VERSION : 0.1
   VAR_INPUT
      digits : String;
   END_VAR
   VAR_TEMP
      _characters : Array[0..#CHAR_COUNT] of Char;
      _count : DInt;
      _i : Int;
      _length : Int;
      _character_count : Int;
      _return : DInt;
      _temp : Bool;
   END_VAR
   VAR CONSTANT
      ASCII_OFFSET : DInt := 16#30;
      BLANK : Time;
      CHAR_COUNT : Int := 9;
      MS_PER_SEC : DInt := 1_000;
   END_VAR
BEGIN
   REGION "EXIT ON NO INPUT"
       IF #digits = '' THEN
           #"Timer.Digits_as_String_to_Seconds" := #BLANK;
           RETURN;
       END_IF;
   END_REGION


   REGION "EXPLODE"
       Strg_TO_Chars(Strg := #digits,
                     pChars := 0,
                     Cnt => #_count,
                     Chars := #_characters);
       #_length := UDINT_TO_INT("Array.Any.Length"(#_characters)) - 1;
   END_REGION


   REGION "COUNT"
       #_character_count := "Array.Char.Search"(array := #_characters, search_term := ' ') - 1;
   END_REGION


   REGION "VALIDATE"
       FOR #_i := 0 TO #_character_count DO
           IF NOT "Char.Is_Numeric"(#_characters[#_i]) THEN
               #"Timer.Digits_as_String_to_Seconds" := #BLANK;
               RETURN;
           END_IF;
       END_FOR;
   END_REGION


   #"Timer.Digits_as_String_to_Seconds" := STRING_TO_DINT(#digits) * #MS_PER_SEC;
END_FUNCTION

FUNCTION "Timer.Digits_as_String_to_Minutes" : Time   // FC267, SCL
{ S7_Optimized_Access := 'TRUE' }
VERSION : 0.1
   VAR_INPUT
      digits : String;
   END_VAR
   VAR CONSTANT
      SECONDS_PER_MINUTE : Int := 60;
   END_VAR
BEGIN
   #"Timer.Digits_as_String_to_Minutes" := #SECONDS_PER_MINUTE * TIME_TO_DINT("Timer.Digits_as_String_to_Seconds"(#digits));
END_FUNCTION

FUNCTION "Timer.Digits_as_String_to_Hours" : Time   // FC269, SCL
{ S7_Optimized_Access := 'TRUE' }
VERSION : 0.1
   VAR_INPUT
      digits : String;
   END_VAR
   VAR CONSTANT
      SECONDS_PER_HOUR : Int := 3_600;
   END_VAR
BEGIN
   #"Timer.Digits_as_String_to_Hours" := #SECONDS_PER_HOUR * TIME_TO_DINT("Timer.Digits_as_String_to_Seconds"(#digits));
END_FUNCTION

// folder: Utilities/UInt

FUNCTION "UInt.Value_Change" : Bool   // FC183, SCL
{ S7_Optimized_Access := 'TRUE' }
VERSION : 0.1
   VAR_INPUT
      value : UInt;
      old_value : UInt;
   END_VAR
BEGIN
   #"UInt.Value_Change" := #value <> #old_value;
END_FUNCTION

// folder: Utilities/USInt

FUNCTION_BLOCK "USInt.State_change"   // FB58, SCL
{ S7_Optimized_Access := 'TRUE' }
VERSION : 0.1
   VAR_INPUT
      value : USInt;
   END_VAR
   VAR_IN_OUT
      get_usint : "State Changes: USInt";
   END_VAR
   VAR
      old_value : USInt;
   END_VAR
   VAR_TEMP
      _return : "State Changes: USInt";
   END_VAR
BEGIN
   REGION "BUFFER IN"
       #_return := #get_usint;
   END_REGION


   REGION "MAP"
       IF #value <> #old_value THEN
           #_return.actual := #value;
       END_IF;
       #_return.rising := "USInt.Rising_Edge"(value := #value,
                                              old_value := #old_value);
       #_return.falling := "USInt.Falling_Edge"(value := #value,
                                                old_value := #old_value);
   END_REGION


   REGION "SAVE OLD VALUE"
       #old_value := #_return.actual;
   END_REGION


   REGION "RETURN" 
       #get_usint := #_return;
   END_REGION
END_FUNCTION_BLOCK

FUNCTION "USInt.Value_Change" : Bool   // FC181, SCL
{ S7_Optimized_Access := 'TRUE' }
VERSION : 0.1
   VAR_INPUT
      value : USInt;
      old_value : USInt;
   END_VAR
BEGIN
   #"USInt.Value_Change" := #value <> #old_value;
END_FUNCTION

FUNCTION "USInt.Rising_Edge" : Bool   // FC262, SCL
{ S7_Optimized_Access := 'TRUE' }
VERSION : 0.1
   VAR_INPUT
      value : USInt;
      old_value : USInt;
   END_VAR
BEGIN
   #"USInt.Rising_Edge" := #value <> "NULL_TOKEN" AND #old_value = "NULL_TOKEN";
END_FUNCTION

FUNCTION "USInt.Falling_Edge" : Bool   // FC263, SCL
{ S7_Optimized_Access := 'TRUE' }
VERSION : 0.1
   VAR_INPUT
      value : USInt;
      old_value : USInt;
   END_VAR
BEGIN
   #"USInt.Falling_Edge" := #value = "NULL_TOKEN" AND #old_value <> "NULL_TOKEN";
END_FUNCTION

// folder: Utilities/WIP

FUNCTION "WIP.Code_to_WString" : WString   // FC64, SCL
{ S7_Optimized_Access := 'TRUE' }
VERSION : 0.1
   VAR_INPUT
      wipTxtLib : "Recipe: Wip Text Library";
      code : DInt;
   END_VAR
   VAR_TEMP
      wipCode : DInt;
      wipText : DInt;
      output : WString;
   END_VAR
   VAR CONSTANT
      newLine : WString := WSTRING#'$L';
   END_VAR
BEGIN
   REGION "PARSE CODE"
       "Part_Number.Parse_Code"(code := #code,
                    code_left => #wipCode,
                    code_right => #wipText);
   END_REGION

   REGION "DOUBLE LINE PN"
       #output := CONCAT_WSTRING(IN1 := #wipTxtLib.code[#wipCode],
                                 IN2 := #newLine,
                                 IN3 := #wipTxtLib.txt[#wipText]);
   END_REGION

   REGION "OUTPUT"
       #"WIP.Code_to_WString" := #output;
   END_REGION
END_FUNCTION

FUNCTION "WIP.Count" : Int   // FC72, SCL
{ S7_Optimized_Access := 'TRUE' }
VERSION : 0.1
   VAR_INPUT
      stnSavedWips : "WIP: Station";
   END_VAR
   VAR_TEMP
      pWip : Int;
   END_VAR
   // Ret_Val : -1 for no wips in station
BEGIN
   WHILE #stnSavedWips.wip[#pWip].wip.code <> -1 DO
       #pWip += 1;
   END_WHILE;
   #"WIP.Count" := #pWip - 1;
END_FUNCTION

FUNCTION "WIP.Global_Index_to_Station" : "WIP: Station"   // FC113, SCL
{ S7_Optimized_Access := 'TRUE' }
VERSION : 0.1
   VAR_INPUT
      index : Int;
      wip_stations : "Recipe: HMI Stations Saved Wips";
   END_VAR
   VAR_TEMP
      i : Int;
      ret : "WIP: Station";
   END_VAR
BEGIN
   REGION "FIND STATION"
       FOR #i := 0 TO "HMI_STATION_COUNT" DO
           IF #wip_stations.stn[#i].pStn = #index THEN
               #ret := #wip_stations.stn[#i];
               EXIT;
           END_IF;
       END_FOR;
   END_REGION


   REGION "RETURN"
       #"WIP.Global_Index_to_Station" := #ret;
   END_REGION
END_FUNCTION

FUNCTION "WIP.Global_Index_to_HMI_Station_Index" : Int   // FC130, SCL
{ S7_Optimized_Access := 'TRUE' }
VERSION : 0.1
   VAR_INPUT
      global_index : Int;
      saved_WIPs : "Recipe: HMI Stations Saved Wips";
   END_VAR
   VAR_TEMP
      i : Int;
      ret : Int;
   END_VAR
BEGIN
   REGION "SEARCH FOR INDEX"
       #ret := "NULL_TOKEN";
       FOR #i := 0 TO "HMI_STATION_COUNT" DO
           IF #saved_WIPs.stn[#i].pStn = #global_index THEN
               #ret := #i;
               EXIT;
           END_IF;
       END_FOR;
   END_REGION


   REGION "RETURN"
       #"WIP.Global_Index_to_HMI_Station_Index" := #ret;
   END_REGION
END_FUNCTION

FUNCTION "WIP.Code_to_Index" : Int   // FC233, SCL
{ S7_Optimized_Access := 'TRUE' }
VERSION : 0.1
   VAR_INPUT
      saved_wip : "WIP: Station";
      wip_code : DInt;
   END_VAR
   VAR_TEMP
      _i : Int;
      _length : Int;
   END_VAR
BEGIN
   #_length := UDINT_TO_INT("Array.Any.Length"(#saved_wip.wip)) - 1;
   FOR #_i := 0 TO #_length DO
       IF #wip_code <> #saved_wip.wip[#_i].wip.code THEN
           CONTINUE;
       END_IF;
       #"WIP.Code_to_Index" := #_i;
       RETURN;
   END_FOR;

   #"WIP.Code_to_Index" := "NULL_TOKEN";
   RETURN;
END_FUNCTION

FUNCTION "WIP_Station.Indices_of_Selected_WIPs" : Void   // FC241, SCL
{ S7_Optimized_Access := 'TRUE' }
VERSION : 0.1
   VAR_INPUT
      selected_wips : "Selected Wips";
      station_wips : "WIP: Station";
   END_VAR
   VAR_IN_OUT
      selected_wip_indices : Array[*] of Int;
   END_VAR
   VAR_TEMP
      _i : Int;
      _length : Int;
      _p_return : Int;
      _wip_index : Int;
   END_VAR
   VAR CONSTANT
      UBOUND : Int := 999;
   END_VAR
BEGIN
   REGION "PREP ARRAY OF FOUND INDICES"
       "Array.Int.Fill"(value := "NULL_TOKEN",
                        int_array := #selected_wip_indices);
       #_length := UDINT_TO_INT("Array.Any.Length"(#selected_wip_indices)) - 1;
   END_REGION

   REGION "FOR EACH SELECTED WIP"
       FOR #_i := 0 TO #selected_wips.count - 1 DO

           REGION "GET SELECTED WIPS INDEX IN THIS STATION"
               #_wip_index := "WIP_Station.Indices_of_Selected_WIPS.Search_WIP"(wip_code := #selected_wips.wips[#_i],
                                                                                station_wips := #station_wips);
           END_REGION

           REGION "IF NOT FOUND GO TO NEXT WIP"
               // fault tolerance
               IF #_wip_index = "NULL_TOKEN" THEN
                   CONTINUE;
               END_IF;
           END_REGION

           REGION "WIP FOUND IN STATION"
               #selected_wip_indices[#_p_return] := #_wip_index;
               #_p_return += 1;
           END_REGION

           REGION "DON'T GO OUT OF FOUND IDEX ARRAY"
               // fault tolerance
               IF #_p_return > #_length THEN
                   RETURN;
               END_IF;
           END_REGION

       END_FOR;
   END_REGION
END_FUNCTION

FUNCTION "WIP_Station.Indices_of_Selected_WIPS.Search_WIP" : Int   // FC242, SCL
{ S7_Optimized_Access := 'TRUE' }
VERSION : 0.1
   VAR_INPUT
      wip_code : DInt;
      station_wips : "WIP: Station";
   END_VAR
   VAR_TEMP
      _i : Int;
      _length : Int;
   END_VAR
BEGIN
   REGION "FOR EACH WIP IN STATION"
       #_length := UDINT_TO_INT("Array.Any.Length"(#station_wips.wip)) - 1;
       FOR #_i := 0 TO #_length DO

           REGION "WIP CODE DOES NOT MATCH"
               IF #wip_code <> #station_wips.wip[#_i].wip.code THEN
                   CONTINUE;
               END_IF;
           END_REGION

           REGION "WIP CODE MATCHES"
               #"WIP_Station.Indices_of_Selected_WIPS.Search_WIP" := #_i;
               RETURN;
           END_REGION

       END_FOR;
   END_REGION

   REGION "NO MATCH FOUND"
       #"WIP_Station.Indices_of_Selected_WIPS.Search_WIP" := "NULL_TOKEN";
       RETURN;
   END_REGION
END_FUNCTION

// folder: Utilities/WString

FUNCTION_BLOCK "WString.State_Change"   // FB51, SCL
{ S7_Optimized_Access := 'TRUE' }
VERSION : 0.1
   VAR_INPUT
      interface : WString;
   END_VAR
   VAR_IN_OUT
      get_wstring : "State Changes: WString";
   END_VAR
   VAR
      old_value : WString;
   END_VAR
   VAR_TEMP
      ret : "State Changes: WString";
   END_VAR
   VAR CONSTANT
      blank : WString;
   END_VAR
BEGIN
   REGION "BUFFER IN"
       #ret := #get_wstring;
   END_REGION


   REGION "MAP"
       IF #interface <> #old_value THEN
           #ret.actual := #interface;
       END_IF;
       #ret.rising := "WString.Rising_Edge"(value := #interface,
                                             old_value := #old_value);
       #ret.falling := "WString.Falling_Edge"(value := #interface,
                                               old_value := #old_value);
   END_REGION


   REGION "SAVE OLD VALUE"
       #old_value := #ret.actual;
   END_REGION


   REGION "RETURN" 
       #get_wstring := #ret;
   END_REGION
END_FUNCTION_BLOCK

FUNCTION "WString.to_Time" : Time   // FC38, SCL
{ S7_Optimized_Access := 'TRUE' }
VERSION : 0.1
   VAR_INPUT
      value : WString;
   END_VAR
   VAR_TEMP
      _component_count : Int;
      _i : Int;
      _return : DInt;
      _time_components : Array[0..4] of WString;
   END_VAR
   VAR CONSTANT
      BLANK : Time;
   END_VAR
BEGIN
   REGION "NO INPUT"
       IF #value = WSTRING#'' THEN
           #"WString.to_Time" := #BLANK;
           RETURN;
       END_IF;
   END_REGION


   REGION "NO DELIMETERS"
       IF FIND(IN1 := WSTRING_TO_STRING(#value), IN2 := ':') = 0 THEN
           IF NOT "WString.to_Time.Validate_Component"(WSTRING_TO_STRING(#value)) THEN
               #"WString.to_Time" := #BLANK;
               RETURN;
           END_IF;
           #_return := "Timer.Digits_as_String_to_Seconds"(WSTRING_TO_STRING(#value));
       END_IF;
   END_REGION


   REGION "EXPLODE INPUT"
       "WString.Split_Single"(wstring_in := #value,
                              delimeter := WString#':',
                              "pointer" := 0,
                              sub_strings := #_time_components);
       #_component_count := "Array.WString.Search"(array := #_time_components, search_term := WString#'') - 1;
   END_REGION


   REGION "EXIT ON TOO MANY COMPONENTS"
       IF #_component_count >= 3 THEN
           #"WString.to_Time" := #BLANK;
       END_IF;
   END_REGION


   REGION "VALIDATE INPUT"
       FOR #_i := 0 TO #_component_count DO
           IF NOT "WString.to_Time.Validate_Component"(WSTRING_TO_STRING(#_time_components[#_i])) THEN
               #"WString.to_Time" := #BLANK;
               RETURN;
           END_IF;
       END_FOR;
   END_REGION


   REGION "REVERSE"
       "Array.WString.Reverse"(null_token := wstring#'',
                               wstring_array := #_time_components);
   END_REGION


   REGION CONVERT ARRAY ELEMENTS TO TIME
       #_return := 0;
       FOR #_i := 0 TO #_component_count DO
           CASE #_i OF
               0:
                   #_return := TIME_TO_DINT("Timer.Digits_as_String_to_Seconds"(WSTRING_TO_STRING(#_time_components[#_i])));
               1:
                   #_return += TIME_TO_DINT("Timer.Digits_as_String_to_Minutes"(WSTRING_TO_STRING(#_time_components[#_i])));
               2:
                   #_return += TIME_TO_DINT("Timer.Digits_as_String_to_Hours"(WSTRING_TO_STRING(#_time_components[#_i])));
           END_CASE;
       END_FOR;
   END_REGION


   REGION RETURN VALUE

       #"WString.to_Time" := DINT_TO_TIME(#_return);

   END_REGION
END_FUNCTION

FUNCTION "WString.Rising_Edge" : Bool   // FC182, SCL
{ S7_Optimized_Access := 'TRUE' }
VERSION : 0.1
   VAR_INPUT
      value : WString;
      old_value : WString;
   END_VAR
   VAR CONSTANT
      blank : WString;
   END_VAR
BEGIN
   #"WString.Rising_Edge" := #value <> #blank AND #old_value = #blank;
END_FUNCTION

FUNCTION "WString.Falling_Edge" : Bool   // FC188, SCL
{ S7_Optimized_Access := 'TRUE' }
VERSION : 0.1
   VAR_INPUT
      value : WString;
      old_value : WString;
   END_VAR
   VAR CONSTANT
      blank : WString;
   END_VAR
BEGIN
   #"WString.Falling_Edge" := #value = #blank AND #old_value <> #blank;
END_FUNCTION

FUNCTION "WString.to_Time.Validate_Component" : Bool   // FC273, SCL
{ S7_Optimized_Access := 'TRUE' }
VERSION : 0.1
   VAR_INPUT
      component : String;
   END_VAR
   VAR_TEMP
      _characters : Array[0..#CHAR_COUNT] of Char;
      _character_count : Int;
      _count : DInt;
      _i : Int;
   END_VAR
   VAR CONSTANT
      CHAR_COUNT : Int := 9;
   END_VAR
BEGIN
   Strg_TO_Chars(Strg := #component,
                 pChars := 0,
                 Cnt => #_count,
                 Chars := #_characters);
   #_character_count := "Array.Char.Search"(array := #_characters, search_term := ' ') - 1;
   FOR #_i := 0 TO #_character_count DO
       IF NOT "Char.Is_Numeric"(#_characters[#_i]) THEN
           #"WString.to_Time.Validate_Component" := FALSE;
           RETURN;
       END_IF;
   END_FOR;
   #"WString.to_Time.Validate_Component" := TRUE;
   RETURN;
END_FUNCTION

// ===== library types =====

TYPE "PB Data"
   STRUCT
      actuate : Bool;
      animate : USInt;
      enable : Bool;
      label : WString[80];
      listSelect : UInt;
      visible : Bool;
   END_STRUCT;
END_TYPE

TYPE "PB Data: Text Label"
   STRUCT
      actuate : Bool;
      animate : USInt;
      label : WString[20];
   END_STRUCT;
END_TYPE

TYPE "Station Assignment: Button Details Data"
   STRUCT
      alloted : Struct
         animate : USInt;
         value : WString[10];
      END_STRUCT;
      critical : Struct
         animate : USInt;
         value : WString[10];
      END_STRUCT;
      label : Struct
         animate : USInt;
         value : WString[2];
      END_STRUCT;
      partNumber : Struct
         animate : USInt;
         value : WString[40];
      END_STRUCT;
      select : Struct
         actuate : Bool;
         animate : USInt;
      END_STRUCT;
   END_STRUCT;
END_TYPE

TYPE "IO Field Data: Timers"
   STRUCT
      animate : USInt;
      inputFinished : Bool;
      value : WString[5];
   END_STRUCT;
END_TYPE

TYPE "Line Label Data"
   STRUCT
      animate : Struct
         bg : USInt;
         ioField : USInt;
      END_STRUCT;
      inputFinished : Bool;
      value : WString[10];
   END_STRUCT;
END_TYPE

TYPE "IO Field Data: Part Number: 2 Line"
   STRUCT
      single_actuate : Bool;
      single_animate : USInt;
      single_enable : Bool;
      single_input_finished : Bool;
      single_value : WString[40];
      single_visible : Bool;
      double_actuate : Bool;
      double_animate : USInt;
      double_enable : Bool;
      double_input_finished_top : Bool;
      double_input_finished_bottom : Bool;
      double_value_top : WString[40];
      double_value_bottom : WString[40];
      double_visible : Bool;
   END_STRUCT;
END_TYPE

TYPE "Drop Zone Data"
   STRUCT
      animate : Struct
         bg : USInt;
         ioField : USInt;
      END_STRUCT;
      inputFinished : Bool;
      value : WString[10];
   END_STRUCT;
END_TYPE

TYPE "Station Sim Data"
   STRUCT
      stn : Struct
         animate : USInt;
         label : WString[20];
      END_STRUCT;
      btn : Struct
         actuate : Byte;
         animate : Array[0..7] of USInt;
         labels : Array[0..7] of WString [4];
      END_STRUCT;
   END_STRUCT;
END_TYPE

// folder: Main HMI

TYPE "Table Row Data"
   STRUCT
      address : DInt := -1;
      ordered : Bool;
      pbSelection : Struct
         actuate : Bool;
         animate : USInt;
      END_STRUCT;
      rtBackground : Struct
         animate : USInt;
      END_STRUCT;
      tfDropZone : Struct
         animate : USInt;
         value : WString[20];
      END_STRUCT;
      tfLine : Struct
         animate : USInt;
         value : WString[20];
      END_STRUCT;
      tfPartNumber : Struct
         animateDL : USInt;
         animateSL : USInt;
         value : WString[40];
      END_STRUCT;
      tfTime : Struct
         animate : USInt;
         value : WString[20];
      END_STRUCT;
   END_STRUCT;
END_TYPE

(* ===== HMI "HMI_RT_1" =====
system functions are stored by id; their names below are inferred from use
connection "Main HMI": ETHERNET, S7_1500_OMS

HMI tags "Default tag table"
   "Clock_Byte" : Byte = PLC Clock_Byte AT %MB0, 100 ms
   "HMI Data: Warehouse HMI_screenNumber" : Int = PLC "HMI Data: Warehouse HMI".screenNumber AT %DB1.DBW0, 100 ms
   "HMI Data: Warehouse HMI_barcode" : Barcode Screen = PLC "HMI Data: Warehouse HMI".barcode AT %DB1.DBW0, 100 ms
   "HMI Data: Warehouse HMI_tableNav_top" : Push Button Data = PLC "HMI Data: Warehouse HMI".tableNav.top, 100 ms
   "HMI Data: Warehouse HMI_tableNav_pageUp" : Push Button Data = PLC "HMI Data: Warehouse HMI".tableNav.pageUp, 100 ms
   "HMI Data: Warehouse HMI_tableNav_lineUp" : Push Button Data = PLC "HMI Data: Warehouse HMI".tableNav.lineUp, 100 ms
   "HMI Data: Warehouse HMI_tableNav_lineDown" : Push Button Data = PLC "HMI Data: Warehouse HMI".tableNav.lineDown, 100 ms
   "HMI Data: Warehouse HMI_tableNav_pageDown" : Push Button Data = PLC "HMI Data: Warehouse HMI".tableNav.pageDown, 100 ms
   "HMI Data: Warehouse HMI_tableNav_bottom" : Push Button Data = PLC "HMI Data: Warehouse HMI".tableNav.bottom, 100 ms
   "HMI Data: Warehouse HMI_networkHealth_pnioDevices{1}" : Push Button Data = PLC "HMI Data: Warehouse HMI".networkHealth.pnioDevices[1], 100 ms
   "HMI Data: Warehouse HMI_networkHealth_pnioDevices{2}" : Push Button Data = PLC "HMI Data: Warehouse HMI".networkHealth.pnioDevices[2], 100 ms
   "HMI Data: Warehouse HMI_networkHealth_pnioDevices{3}" : Push Button Data = PLC "HMI Data: Warehouse HMI".networkHealth.pnioDevices[3], 100 ms
   "HMI Data: Warehouse HMI_networkHealth_pnioDevices{4}" : Push Button Data = PLC "HMI Data: Warehouse HMI".networkHealth.pnioDevices[4], 100 ms
   "HMI Data: Warehouse HMI_networkHealth_pnioDevices{5}" : Push Button Data = PLC "HMI Data: Warehouse HMI".networkHealth.pnioDevices[5], 100 ms
   "HMI Data: Warehouse HMI_networkHealth_pnioDevices{6}" : Push Button Data = PLC "HMI Data: Warehouse HMI".networkHealth.pnioDevices[6], 100 ms
   "HMI Data: Warehouse HMI_networkHealth_pnioDevices{7}" : Push Button Data = PLC "HMI Data: Warehouse HMI".networkHealth.pnioDevices[7], 100 ms
   "HMI Data: Warehouse HMI_networkHealth_pnioDevices{8}" : Push Button Data = PLC "HMI Data: Warehouse HMI".networkHealth.pnioDevices[8], 100 ms
   "HMI Data: Warehouse HMI_networkHealth_pnioDevices{9}" : Push Button Data = PLC "HMI Data: Warehouse HMI".settings.selectStation, 100 ms
   "HMI Data: Warehouse HMI_networkHealth_pnioDevices{10}" : Push Button Data = PLC "HMI Data: Warehouse HMI".networkHealth.pnioDevices[10], 100 ms
   "HMI Data: Warehouse HMI_networkHealth_pnioDevices{11}" : Push Button Data = PLC "HMI Data: Warehouse HMI".networkHealth.pnioDevices[11], 100 ms
   "HMI Data: Warehouse HMI_networkHealth_pnioDevices{12}" : Push Button Data = PLC "HMI Data: Warehouse HMI".networkHealth.pnioDevices[12], 100 ms
   "HMI Data: Warehouse HMI_networkHealth_pnioDevices{13}" : Push Button Data = PLC "HMI Data: Warehouse HMI".networkHealth.pnioDevices[13], 100 ms
   "HMI Data: Warehouse HMI_networkHealth_pnioDevices{16}" : Push Button Data = PLC "HMI Data: Warehouse HMI".networkHealth.pnioDevices[16], 100 ms
   "HMI Data: Warehouse HMI_networkHealth_pnioDevices{14}" : Push Button Data = PLC "HMI Data: Warehouse HMI".networkHealth.pnioDevices[14], 100 ms
   "HMI Data: Warehouse HMI_networkHealth_pnioDevices{15}" : Push Button Data = PLC "HMI Data: Warehouse HMI".networkHealth.pnioDevices[15], 100 ms
   "HMI Data: Warehouse HMI_networkHealth_pnioDevices{17}" : Push Button Data = PLC "HMI Data: Warehouse HMI".networkHealth.pnioDevices[17], 100 ms
   "HMI Data: Warehouse HMI_networkHealth_pnioDevices{18}" : Push Button Data = PLC "HMI Data: Warehouse HMI".networkHealth.pnioDevices[18], 100 ms
   "HMI Data: Warehouse HMI_networkHealth_pnioDevices{19}" : Push Button Data = PLC "HMI Data: Warehouse HMI".networkHealth.pnioDevices[19], 100 ms
   "HMI Data: Warehouse HMI_networkHealth_pnioDevices{20}" : Push Button Data = PLC "HMI Data: Warehouse HMI".networkHealth.pnioDevices[20], 100 ms
   "HMI Data: Warehouse HMI_networkHealth_pnioDevices{21}" : Push Button Data = PLC "HMI Data: Warehouse HMI".networkHealth.pnioDevices[21], 100 ms
   "HMI Data: Warehouse HMI_networkHealth_pnioDevices{22}" : Push Button Data = PLC "HMI Data: Warehouse HMI".networkHealth.pnioDevices[22], 100 ms
   "HMI Data: Warehouse HMI_networkHealth_pnioDevices{31}" : Push Button Data = PLC "HMI Data: Warehouse HMI".networkHealth.pnioDevices[31], 100 ms
   "HMI Data: Warehouse HMI_networkHealth_pnioDevices{32}" : Push Button Data = PLC "HMI Data: Warehouse HMI".networkHealth.pnioDevices[32], 100 ms
   "HMI Data: Warehouse HMI_networkHealth_pnioDevices{29}" : Push Button Data = PLC "HMI Data: Warehouse HMI".networkHealth.pnioDevices[29], 100 ms
   "HMI Data: Warehouse HMI_networkHealth_pnioDevices{30}" : Push Button Data = PLC "HMI Data: Warehouse HMI".networkHealth.pnioDevices[30], 100 ms
   "HMI Data: Warehouse HMI_networkHealth_pnioDevices{27}" : Push Button Data = PLC "HMI Data: Warehouse HMI".networkHealth.pnioDevices[27], 100 ms
   "HMI Data: Warehouse HMI_networkHealth_pnioDevices{28}" : Push Button Data = PLC "HMI Data: Warehouse HMI".networkHealth.pnioDevices[28], 100 ms
   "HMI Data: Warehouse HMI_networkHealth_pnioDevices{23}" : Push Button Data = PLC "HMI Data: Warehouse HMI".networkHealth.pnioDevices[23], 100 ms
   "HMI Data: Warehouse HMI_networkHealth_pnioDevices{24}" : Push Button Data = PLC "HMI Data: Warehouse HMI".networkHealth.pnioDevices[24], 100 ms
   "HMI Data: Warehouse HMI_networkHealth_pnioDevices{25}" : Push Button Data = PLC "HMI Data: Warehouse HMI".networkHealth.pnioDevices[25], 100 ms
   "HMI Data: Warehouse HMI_networkHealth_pnioDevices{26}" : Push Button Data = PLC "HMI Data: Warehouse HMI".networkHealth.pnioDevices[26], 100 ms
   "HMI Data: Warehouse HMI_networkHealth_pnioDevices{33}" : Push Button Data = PLC "HMI Data: Warehouse HMI".networkHealth.pnioDevices[33], 100 ms
   "HMI Data: Warehouse HMI_networkHealth_pnioDevices{34}" : Push Button Data = PLC "HMI Data: Warehouse HMI".networkHealth.pnioDevices[34], 100 ms
   "HMI Data: Warehouse HMI_networkHealth_pnioDevices{35}" : Push Button Data = PLC "HMI Data: Warehouse HMI".networkHealth.pnioDevices[35], 100 ms
   "HMI Data: Warehouse HMI_networkHealth_pnioDevices{36}" : Push Button Data = PLC "HMI Data: Warehouse HMI".networkHealth.pnioDevices[36], 100 ms
   "HMI Data: Warehouse HMI_networkHealth_pnioDevices{37}" : Push Button Data = PLC "HMI Data: Warehouse HMI".networkHealth.pnioDevices[37], 100 ms
   "HMI Data: Warehouse HMI_networkHealth_pnioDevices{38}" : Push Button Data = PLC "HMI Data: Warehouse HMI".networkHealth.pnioDevices[38], 100 ms
   "HMI Data: Warehouse HMI_networkHealth_pnioDevices{39}" : Push Button Data = PLC "HMI Data: Warehouse HMI".networkHealth.pnioDevices[39], 100 ms
   "HMI Data: Warehouse HMI_networkHealth_pnioDevices{40}" : Push Button Data = PLC "HMI Data: Warehouse HMI".networkHealth.pnioDevices[40], 100 ms
   "HMI Data: Warehouse HMI_networkHealth_pnioDevices{41}" : Push Button Data = PLC "HMI Data: Warehouse HMI".networkHealth.pnioDevices[41], 100 ms
   "HMI Data: Warehouse HMI_networkHealth_pnioDevices{42}" : Push Button Data = PLC "HMI Data: Warehouse HMI".networkHealth.pnioDevices[42], 100 ms
   "HMI Data: Warehouse HMI_networkHealth_pnioDevices{43}" : Push Button Data = PLC "HMI Data: Warehouse HMI".networkHealth.pnioDevices[43], 100 ms
   "HMI Data: Warehouse HMI_networkHealth_pnioDevices{44}" : Push Button Data = PLC "HMI Data: Warehouse HMI".networkHealth.pnioDevices[44], 100 ms
   "HMI Data: Warehouse HMI_networkHealth_pnioDevices{45}" : Push Button Data = PLC "HMI Data: Warehouse HMI".networkHealth.pnioDevices[45], 100 ms
   "HMI Data: Warehouse HMI_networkHealth_pnioDevices{46}" : Push Button Data = PLC "HMI Data: Warehouse HMI".networkHealth.pnioDevices[46], 100 ms
   "HMI Data: Warehouse HMI_networkHealth_pnioDevices{47}" : Push Button Data = PLC "HMI Data: Warehouse HMI".networkHealth.pnioDevices[47], 100 ms
   "HMI Data: Warehouse HMI_networkHealth_pnioDevices{48}" : Push Button Data = PLC "HMI Data: Warehouse HMI".networkHealth.pnioDevices[48], 100 ms
   "HMI Data: Warehouse HMI_networkHealth_et200spPopUp" : Station: ET200SP Comm Debug Data = PLC "HMI Data: Warehouse HMI".networkHealth.et200spPopUp, 100 ms
   "HMI Data: Warehouse HMI_networkHealth_kp8PopUp" : Station: KP8 Comm Debug Data = PLC "HMI Data: Warehouse HMI".networkHealth.kp8PopUp, 100 ms
   "HMI Data: Warehouse HMI_networkHealth_selectedDevice" : Int = PLC "HMI Data: Warehouse HMI".networkHealth.selectedDevice, 100 ms

HMI tags "Pop Ups: Select Buttons"
   "HMI Data: Warehouse HMI_pop_up_select_buttons_buttons{0}" : Push Button Data = PLC "HMI Data: Warehouse HMI".pop_up.select_buttons.buttons[0], 100 ms
   "HMI Data: Warehouse HMI_pop_up_select_buttons_buttons{1}" : Push Button Data = PLC "HMI Data: Warehouse HMI".pop_up.select_buttons.buttons[1], 100 ms
   "HMI Data: Warehouse HMI_pop_up_select_buttons_buttons{2}" : Push Button Data = PLC "HMI Data: Warehouse HMI".pop_up.select_buttons.buttons[2], 100 ms
   "HMI Data: Warehouse HMI_pop_up_select_buttons_buttons{3}" : Push Button Data = PLC "HMI Data: Warehouse HMI".pop_up.select_buttons.buttons[3], 100 ms
   "HMI Data: Warehouse HMI_pop_up_select_buttons_buttons{4}" : Push Button Data = PLC "HMI Data: Warehouse HMI".pop_up.select_buttons.buttons[4], 100 ms
   "HMI Data: Warehouse HMI_pop_up_select_buttons_buttons{5}" : Push Button Data = PLC "HMI Data: Warehouse HMI".pop_up.select_buttons.buttons[5], 100 ms
   "HMI Data: Warehouse HMI_pop_up_select_buttons_buttons{6}" : Push Button Data = PLC "HMI Data: Warehouse HMI".pop_up.select_buttons.buttons[6], 100 ms
   "HMI Data: Warehouse HMI_pop_up_select_buttons_buttons{7}" : Push Button Data = PLC "HMI Data: Warehouse HMI".pop_up.select_buttons.buttons[7], 100 ms
   "HMI Data: Warehouse HMI_pop_up_select_buttons_close_screen" : Push Button Data = PLC "HMI Data: Warehouse HMI".pop_up.select_buttons.close_screen, 100 ms

HMI tags "Pop Ups: Select Stations"
   "HMI Data: Warehouse HMI_pop_up_select_stations_close_screen" : Push Button Data = PLC "HMI Data: Warehouse HMI".pop_up.select_stations.close_screen, 100 ms
   "HMI Data: Warehouse HMI_pop_up_select_stations_nav_bar_hmi" : Nav Bar Data: HMI = PLC "HMI Data: Warehouse HMI".pop_up.select_stations.nav_bar.hmi, 100 ms
   "HMI Data: Warehouse HMI_pop_up_select_stations_stn_select_btns{0}" : Push Button Data = PLC "HMI Data: Warehouse HMI".pop_up.select_stations.stn_select_btns[0], 100 ms
   "HMI Data: Warehouse HMI_pop_up_select_stations_stn_select_btns{1}" : Push Button Data = PLC "HMI Data: Warehouse HMI".pop_up.select_stations.stn_select_btns[1], 100 ms
   "HMI Data: Warehouse HMI_pop_up_select_stations_stn_select_btns{10}" : Push Button Data = PLC "HMI Data: Warehouse HMI".pop_up.select_stations.stn_select_btns[10], 100 ms
   "HMI Data: Warehouse HMI_pop_up_select_stations_stn_select_btns{11}" : Push Button Data = PLC "HMI Data: Warehouse HMI".pop_up.select_stations.stn_select_btns[11], 100 ms
   "HMI Data: Warehouse HMI_pop_up_select_stations_stn_select_btns{2}" : Push Button Data = PLC "HMI Data: Warehouse HMI".pop_up.select_stations.stn_select_btns[2], 100 ms
   "HMI Data: Warehouse HMI_pop_up_select_stations_stn_select_btns{3}" : Push Button Data = PLC "HMI Data: Warehouse HMI".pop_up.select_stations.stn_select_btns[3], 100 ms
   "HMI Data: Warehouse HMI_pop_up_select_stations_stn_select_btns{4}" : Push Button Data = PLC "HMI Data: Warehouse HMI".pop_up.select_stations.stn_select_btns[4], 100 ms
   "HMI Data: Warehouse HMI_pop_up_select_stations_stn_select_btns{5}" : Push Button Data = PLC "HMI Data: Warehouse HMI".pop_up.select_stations.stn_select_btns[5], 100 ms
   "HMI Data: Warehouse HMI_pop_up_select_stations_stn_select_btns{6}" : Push Button Data = PLC "HMI Data: Warehouse HMI".pop_up.select_stations.stn_select_btns[6], 100 ms
   "HMI Data: Warehouse HMI_pop_up_select_stations_stn_select_btns{7}" : Push Button Data = PLC "HMI Data: Warehouse HMI".pop_up.select_stations.stn_select_btns[7], 100 ms
   "HMI Data: Warehouse HMI_pop_up_select_stations_stn_select_btns{8}" : Push Button Data = PLC "HMI Data: Warehouse HMI".pop_up.select_stations.stn_select_btns[8], 100 ms
   "HMI Data: Warehouse HMI_pop_up_select_stations_stn_select_btns{9}" : Push Button Data = PLC "HMI Data: Warehouse HMI".pop_up.select_stations.stn_select_btns[9], 100 ms

HMI tags "Pop Ups: Select WIPs"
   "HMI Data: Warehouse HMI_pop_up_select_WIPs_select_wip_buttons{0}" : Push Button Data = PLC "HMI Data: Warehouse HMI".pop_up.select_WIPs.select_wip_buttons[0], 100 ms
   "HMI Data: Warehouse HMI_pop_up_select_WIPs_select_wip_buttons{1}" : Push Button Data = PLC "HMI Data: Warehouse HMI".pop_up.select_WIPs.select_wip_buttons[1], 100 ms
   "HMI Data: Warehouse HMI_pop_up_select_WIPs_select_wip_buttons{2}" : Push Button Data = PLC "HMI Data: Warehouse HMI".pop_up.select_WIPs.select_wip_buttons[2], 100 ms
   "HMI Data: Warehouse HMI_pop_up_select_WIPs_select_wip_buttons{3}" : Push Button Data = PLC "HMI Data: Warehouse HMI".pop_up.select_WIPs.select_wip_buttons[3], 100 ms
   "HMI Data: Warehouse HMI_pop_up_select_WIPs_select_wip_buttons{4}" : Push Button Data = PLC "HMI Data: Warehouse HMI".pop_up.select_WIPs.select_wip_buttons[4], 100 ms
   "HMI Data: Warehouse HMI_pop_up_select_WIPs_select_wip_buttons{5}" : Push Button Data = PLC "HMI Data: Warehouse HMI".pop_up.select_WIPs.select_wip_buttons[5], 100 ms
   "HMI Data: Warehouse HMI_pop_up_select_WIPs_select_wip_buttons{6}" : Push Button Data = PLC "HMI Data: Warehouse HMI".pop_up.select_WIPs.select_wip_buttons[6], 100 ms
   "HMI Data: Warehouse HMI_pop_up_select_WIPs_close_screen" : Push Button Data = PLC "HMI Data: Warehouse HMI".pop_up.select_WIPs.close_screen, 100 ms
   "HMI Data: Warehouse HMI_pop_up_select_WIPs_nav_bar_hmi" : Nav Bar Data: HMI = PLC "HMI Data: Warehouse HMI".pop_up.select_WIPs.nav_bar.hmi, 100 ms

HMI tags "Part Call"
   "HMI Data: Warehouse HMI_partCall_row{0}" : Table Row = PLC "HMI Data: Warehouse HMI".partCall.row[0], 100 ms
   "HMI Data: Warehouse HMI_partCall_row{1}" : Table Row = PLC "HMI Data: Warehouse HMI".partCall.row[1], 100 ms
   "HMI Data: Warehouse HMI_partCall_row{10}" : Table Row = PLC "HMI Data: Warehouse HMI".partCall.row[10], 100 ms
   "HMI Data: Warehouse HMI_partCall_row{2}" : Table Row = PLC "HMI Data: Warehouse HMI".partCall.row[2], 100 ms
   "HMI Data: Warehouse HMI_partCall_row{3}" : Table Row = PLC "HMI Data: Warehouse HMI".partCall.row[3], 100 ms
   "HMI Data: Warehouse HMI_partCall_row{4}" : Table Row = PLC "HMI Data: Warehouse HMI".partCall.row[4], 100 ms
   "HMI Data: Warehouse HMI_partCall_row{5}" : Table Row = PLC "HMI Data: Warehouse HMI".partCall.row[5], 100 ms
   "HMI Data: Warehouse HMI_partCall_row{6}" : Table Row = PLC "HMI Data: Warehouse HMI".partCall.row[6], 100 ms
   "HMI Data: Warehouse HMI_partCall_row{7}" : Table Row = PLC "HMI Data: Warehouse HMI".partCall.row[7], 100 ms
   "HMI Data: Warehouse HMI_partCall_row{8}" : Table Row = PLC "HMI Data: Warehouse HMI".partCall.row[8], 100 ms
   "HMI Data: Warehouse HMI_partCall_row{9}" : Table Row = PLC "HMI Data: Warehouse HMI".partCall.row[9], 100 ms

HMI tags "Sim Stations"
   "HMI Data: Warehouse HMI_simStations_down" : Push Button Data = PLC "HMI Data: Warehouse HMI".simStations.down, 100 ms
   "HMI Data: Warehouse HMI_simStations_me{0}" : Station: Sim Data = PLC "HMI Data: Warehouse HMI".simStations.me[0] AT %DB1.DBX0.0, 100 ms
   "HMI Data: Warehouse HMI_simStations_me{1}" : Station: Sim Data = PLC "HMI Data: Warehouse HMI".simStations.me[1], 100 ms
   "HMI Data: Warehouse HMI_simStations_me{10}" : Station: Sim Data = PLC "HMI Data: Warehouse HMI".simStations.me[10], 100 ms
   "HMI Data: Warehouse HMI_simStations_me{11}" : Station: Sim Data = PLC "HMI Data: Warehouse HMI".simStations.me[11], 100 ms
   "HMI Data: Warehouse HMI_simStations_me{2}" : Station: Sim Data = PLC "HMI Data: Warehouse HMI".simStations.me[2], 100 ms
   "HMI Data: Warehouse HMI_simStations_me{3}" : Station: Sim Data = PLC "HMI Data: Warehouse HMI".simStations.me[3], 100 ms
   "HMI Data: Warehouse HMI_simStations_me{4}" : Station: Sim Data = PLC "HMI Data: Warehouse HMI".simStations.me[4], 100 ms
   "HMI Data: Warehouse HMI_simStations_me{5}" : Station: Sim Data = PLC "HMI Data: Warehouse HMI".simStations.me[5], 100 ms
   "HMI Data: Warehouse HMI_simStations_me{6}" : Station: Sim Data = PLC "HMI Data: Warehouse HMI".simStations.me[6], 100 ms
   "HMI Data: Warehouse HMI_simStations_me{7}" : Station: Sim Data = PLC "HMI Data: Warehouse HMI".simStations.me[7], 100 ms
   "HMI Data: Warehouse HMI_simStations_me{8}" : Station: Sim Data = PLC "HMI Data: Warehouse HMI".simStations.me[8], 100 ms
   "HMI Data: Warehouse HMI_simStations_me{9}" : Station: Sim Data = PLC "HMI Data: Warehouse HMI".simStations.me[9], 100 ms
   "HMI Data: Warehouse HMI_simStations_up" : Push Button Data = PLC "HMI Data: Warehouse HMI".simStations.up, 100 ms

HMI tags "Settings: Interface"
   "HMI Data: Warehouse HMI_settings_assign" : Push Button Data = PLC "HMI Data: Warehouse HMI".settings.assign, 100 ms
   "HMI Data: Warehouse HMI_settings_partNumber" : Part_Number_Double.UDT = PLC "HMI Data: Warehouse HMI".settings.partNumber, 100 ms
   "HMI Data: Warehouse HMI_settings_critical" : IO Field Data: Label with Data = PLC "HMI Data: Warehouse HMI".settings.critical, 100 ms
   "HMI Data: Warehouse HMI_settings_total" : IO Field Data: Label with Data = PLC "HMI Data: Warehouse HMI".settings.total, 100 ms
   "HMI Data: Warehouse HMI_settings_dropzone" : IO Field Data: Label with Data = PLC "HMI Data: Warehouse HMI".settings.dropzone, 100 ms
   "HMI Data: Warehouse HMI_settings_line" : IO Field Data: Label with Data = PLC "HMI Data: Warehouse HMI".settings.line, 100 ms
   "HMI Data: Warehouse HMI_settings_selectButton" : Push Button Data = PLC "HMI Data: Warehouse HMI".settings.selectButton, 100 ms
   "HMI Data: Warehouse HMI_settings_selectWip" : Push Button Data = PLC "HMI Data: Warehouse HMI".settings.selectWip, 100 ms
   "HMI Data: Warehouse HMI_settings_selectStation" : Push Button Data = PLC "HMI Data: Warehouse HMI".settings.selectStation, 100 ms
   "HMI Data: Warehouse HMI_settings_stnTableNavBar_hmi" : Nav Bar Data: HMI = PLC "HMI Data: Warehouse HMI".settings.stnTableNavBar.hmi AT %DB1.DBW0, 100 ms

HMI tags "Settings: Feedback"
   "HMI Data: Warehouse HMI_settings_stationRows{0}" : Settings Station Row Data = PLC "HMI Data: Warehouse HMI".settings.stationRows[0], 100 ms
   "HMI Data: Warehouse HMI_settings_stationRows{1}" : Settings Station Row Data = PLC "HMI Data: Warehouse HMI".settings.stationRows[1], 100 ms
   "HMI Data: Warehouse HMI_settings_stationRows{2}" : Settings Station Row Data = PLC "HMI Data: Warehouse HMI".settings.stationRows[2], 100 ms

graphic list "Vertical Table Nav Bar": 0 '100 x 100 Top'; 1 '100 x 100 Actuated Top'; 2 '100 x 100 Page Up'; 3 '100 x 100 Actuated Page Up'; 4 '100 x 100 Line Up'; 5 '100 x 100 Actuated Line Up'; 6 '100 x 100 Line Down'; 7 '100 x 100 Actuated Line Down'; 8 '100 x 100 Page Down'; 9 '100 x 100 Actuated Page Down'; 10 '100 x 100 Bottom'; 11 '100 x 100 Actuated Bottom'

screen "1 PART CALL" 1366x768
   on GenerateScreen: SetTag("HMI Data: Warehouse HMI_screenNumber", 1)
   Rectangle "Settings Tab Background" at 682,0 size 684x68
      Appearance <- "HMI Data: Warehouse HMI_screenNumber"
   Rectangle "Part Call Tab Background" at 0,0 size 685x68
      Appearance <- "HMI Data: Warehouse HMI_screenNumber"
   Rectangle "Settings Tab Border Hide" at 685,61 size 678x20
      Visibility <- "HMI Data: Warehouse HMI_screenNumber"
   Rectangle "Part Call Tab Border Hide" at 3,61 size 679x20
      Visibility <- "HMI Data: Warehouse HMI_screenNumber"
   Button "Settings Screen" at 683,0 size 683x68; TextOff 'SETTINGS'; Authorization "User administration"
      on Release: ActivateScreen("2 SETTINGS", 0)
   Button "Part Call Screen" at 0,0 size 683x68; TextOff 'PART CALL'
      on Release: ActivateScreen("1 PART CALL", 0)
   TextField "Header Line" at 32,112 size 216x53; Text 'LINE'
   TextField "Header Drop Zone" at 238,112 size 236x53; Text 'DROP ZONE'
   TextField "Header Part Number" at 474,112 size 648x53; Text 'PART NUMBER'
   TextField "Header Time" at 1112,112 size 222x53; Text 'TIME'
   ScreenModuleView "TableRow00" at 27,170 size 1312x52; ScreenModuleType ""
      Guid_{11997190-27688} <- "HMI Data: Warehouse HMI_partCall_row{0}"
      on Guid_{11997190-83214}: ActivateScreen("3 BARCODE", 0)
   ScreenModuleView "TableRow01" at 27,222 size 1312x52; ScreenModuleType ""
      Guid_{11997190-27688} <- "HMI Data: Warehouse HMI_partCall_row{1}"
      on Guid_{11997190-83214}: ActivateScreen("3 BARCODE", 0)
   ScreenModuleView "TableRow02" at 27,274 size 1312x52; ScreenModuleType ""
      Guid_{11997190-27688} <- "HMI Data: Warehouse HMI_partCall_row{2}"
      on Guid_{11997190-83214}: ActivateScreen("3 BARCODE", 0)
   ScreenModuleView "TableRow03" at 27,326 size 1312x52; ScreenModuleType ""
      Guid_{11997190-27688} <- "HMI Data: Warehouse HMI_partCall_row{3}"
      on Guid_{11997190-83214}: ActivateScreen("3 BARCODE", 0)
   ScreenModuleView "TableRow04" at 27,378 size 1312x52; ScreenModuleType ""
      Guid_{11997190-27688} <- "HMI Data: Warehouse HMI_partCall_row{4}"
      on Guid_{11997190-83214}: ActivateScreen("3 BARCODE", 0)
   ScreenModuleView "TableRow05" at 27,430 size 1312x52; ScreenModuleType ""
      Guid_{11997190-27688} <- "HMI Data: Warehouse HMI_partCall_row{5}"
      on Guid_{11997190-83214}: ActivateScreen("3 BARCODE", 0)
   ScreenModuleView "TableRow06" at 27,482 size 1312x52; ScreenModuleType ""
      Guid_{11997190-27688} <- "HMI Data: Warehouse HMI_partCall_row{6}"
      on Guid_{11997190-83214}: ActivateScreen("3 BARCODE", 0)
   ScreenModuleView "TableRow07" at 27,534 size 1312x52; ScreenModuleType ""
      Guid_{11997190-27688} <- "HMI Data: Warehouse HMI_partCall_row{7}"
      on Guid_{11997190-83214}: ActivateScreen("3 BARCODE", 0)
   ScreenModuleView "TableRow08" at 27,586 size 1312x52; ScreenModuleType ""
      Guid_{11997190-27688} <- "HMI Data: Warehouse HMI_partCall_row{8}"
      on Guid_{11997190-83214}: ActivateScreen("3 BARCODE", 0)
   ScreenModuleView "TableRow09" at 27,638 size 1312x52; ScreenModuleType ""
      Guid_{11997190-27688} <- "HMI Data: Warehouse HMI_partCall_row{9}"
      on Guid_{11997190-83214}: ActivateScreen("3 BARCODE", 0)
   ScreenModuleView "TableRow10" at 27,690 size 1312x52; ScreenModuleType ""
      Guid_{11997190-27688} <- "HMI Data: Warehouse HMI_partCall_row{10}"
      on Guid_{11997190-83214}: ActivateScreen("3 BARCODE", 0)

SlideinScreen "GraphX_Slidein_Bottom" 1366x80
   ScreenModuleView "Top" at 0,0 size 227x80; Guid_{11997190-63799} "Top"; ScreenModuleType ""
      Guid_{11997190-63779} <- "HMI Data: Warehouse HMI_tableNav_top"
   ScreenModuleView "Page Up" at 227,0 size 228x80; Guid_{11997190-63799} "pageUp"; ScreenModuleType ""
      Guid_{11997190-63779} <- "HMI Data: Warehouse HMI_tableNav_pageUp"
   ScreenModuleView "Line Up" at 455,0 size 228x80; Guid_{11997190-63799} "Up"; ScreenModuleType ""
      Guid_{11997190-63779} <- "HMI Data: Warehouse HMI_tableNav_lineUp"
   ScreenModuleView "Line Down" at 683,0 size 228x80; Guid_{11997190-63799} "Down"; ScreenModuleType ""
      Guid_{11997190-63779} <- "HMI Data: Warehouse HMI_tableNav_lineDown"
   ScreenModuleView "Page Down" at 911,0 size 228x80; Guid_{11997190-63799} "PageDown"; ScreenModuleType ""
      Guid_{11997190-63779} <- "HMI Data: Warehouse HMI_tableNav_pageDown"
   ScreenModuleView "Bottom" at 1138,0 size 228x80; Guid_{11997190-63799} "Bottom"; ScreenModuleType ""
      Guid_{11997190-63779} <- "HMI Data: Warehouse HMI_tableNav_bottom"
   TextField "Text field_1" at 0,0 size 1366x80; Text 'NOT USED'
      Visibility <- "HMI Data: Warehouse HMI_screenNumber"

SlideinScreen "GraphX_Slidein_Right" 449x768
   ScreenModuleView "Station Sim_1" at 5,5 size 106x232; ScreenModuleType ""
      Guid_{11997190-89108} <- "HMI Data: Warehouse HMI_simStations_me{0}"
   ScreenModuleView "Station Sim_2" at 116,5 size 106x232; ScreenModuleType ""
      Guid_{11997190-89108} <- "HMI Data: Warehouse HMI_simStations_me{1}"
   ScreenModuleView "Station Sim_3" at 227,5 size 106x232; ScreenModuleType ""
      Guid_{11997190-89108} <- "HMI Data: Warehouse HMI_simStations_me{2}"
   ScreenModuleView "Station Sim_4" at 338,5 size 106x232; ScreenModuleType ""
      Guid_{11997190-89108} <- "HMI Data: Warehouse HMI_simStations_me{3}"
   ScreenModuleView "Station Sim_5" at 5,242 size 106x232; ScreenModuleType ""
      Guid_{11997190-89108} <- "HMI Data: Warehouse HMI_simStations_me{4}"
   ScreenModuleView "Station Sim_6" at 5,479 size 106x232; ScreenModuleType ""
      Guid_{11997190-89108} <- "HMI Data: Warehouse HMI_simStations_me{8}"
   ScreenModuleView "Station Sim_7" at 116,242 size 106x232; ScreenModuleType ""
      Guid_{11997190-89108} <- "HMI Data: Warehouse HMI_simStations_me{5}"
   ScreenModuleView "Station Sim_8" at 227,242 size 106x232; ScreenModuleType ""
      Guid_{11997190-89108} <- "HMI Data: Warehouse HMI_simStations_me{6}"
   ScreenModuleView "Station Sim_9" at 338,242 size 106x232; ScreenModuleType ""
      Guid_{11997190-89108} <- "HMI Data: Warehouse HMI_simStations_me{7}"
   ScreenModuleView "Station Sim_10" at 116,479 size 106x232; ScreenModuleType ""
      Guid_{11997190-89108} <- "HMI Data: Warehouse HMI_simStations_me{9}"
   ScreenModuleView "Station Sim_11" at 227,478 size 106x232; ScreenModuleType ""
      Guid_{11997190-89108} <- "HMI Data: Warehouse HMI_simStations_me{10}"
   ScreenModuleView "Station Sim_12" at 338,477 size 106x232; ScreenModuleType ""
      Guid_{11997190-89108} <- "HMI Data: Warehouse HMI_simStations_me{11}"
   ScreenModuleView "PB: Graphic/Text List_1" at 5,716 size 65x45; Guid_{11997190-63799} "Up"; ScreenModuleType ""
      Guid_{11997190-63779} <- "HMI Data: Warehouse HMI_simStations_up"
   ScreenModuleView "PB: Graphic/Text List_2" at 379,716 size 65x45; Guid_{11997190-63799} "Down"; ScreenModuleType ""
      Guid_{11997190-63779} <- "HMI Data: Warehouse HMI_simStations_down"

screen "3 BARCODE" 1366x768
   on GenerateScreen: SetTag("HMI Data: Warehouse HMI_screenNumber", 3)
   Rectangle "Nav Panel 02" at 682,700 size 684x68
      Appearance <- "HMI Data: Warehouse HMI_screenNumber"
   Rectangle "Nav Panel 01" at 0,700 size 685x68
      Appearance <- "HMI Data: Warehouse HMI_screenNumber"
   Rectangle "Nav Panel 03 Top Border Hide" at 685,700 size 678x3
      Visibility <- "HMI Data: Warehouse HMI_screenNumber"
   Rectangle "Nav Panel 01 Top Border Hide" at 3,700 size 679x3
      Visibility <- "HMI Data: Warehouse HMI_screenNumber"
   Button "Settings Screen" at 683,700 size 683x68; TextOff 'SETTINGS'; Authorization "User administration"
      on Release: ActivateScreen("2 SETTINGS", 0)
   Button "Part Call Screen" at 0,700 size 683x68; TextOff 'PART CALL'
      on Release: ActivateScreen("1 PART CALL", 0)
   Button "btCancel" at 685,431 size 649x68; TextOff 'CANCEL'
      on Release: ActivateScreen("1 PART CALL", 0)
   Button "btPartOrdered" at 32,431 size 648x68; TextOff 'ORDERED'
      on Release: SetBit("ordered"); ActivateScreen("1 PART CALL", 0)
   TextField "tfBarcodeDisplay" at 32,220 size 1302x206; Text 'Text'
   TextField "tfPartNumberDisplay" at 32,160 size 1302x53; Text 'BARCODE FOR PART NUMBER'

PopupScreen "KP8 Comm Status" 438x720
   ScreenModuleView "Station: KP8_1" at 5,5 size 428x710; ScreenModuleType ""
      Guid_{11997190-107144} <- "HMI Data: Warehouse HMI_networkHealth_kp8PopUp"
      on Guid_{11997190-107182}: function_efd93a16("KP8 Comm Status", 0, 0, -1, -1, 1)

PopupScreen "ET200SP Comm Status" 613x720
   ScreenModuleView "Station: ET200SP_1" at 5,5 size 603x710; ScreenModuleType ""
      Guid_{11997190-102952} <- "HMI Data: Warehouse HMI_networkHealth_et200spPopUp"
      on Guid_{11997190-102950}: function_efd93a16("ET200SP Comm Status", 0, 0, -1, -1, 1)

screen "2 SETTINGS" 1366x768
   on GenerateScreen: SetTag("HMI Data: Warehouse HMI_screenNumber", 2)
   Rectangle "Part Call Nave Panel" at 0,0 size 455x68
      Appearance <- "HMI Data: Warehouse HMI_screenNumber"
   Rectangle "Settings Nav Panel" at 452,0 size 462x68
      Appearance <- "HMI Data: Warehouse HMI_screenNumber"
   Rectangle "Network Health Nav Panel" at 911,0 size 455x68
      Appearance <- "HMI Data: Warehouse HMI_screenNumber"
   Rectangle "Part Call Border Hide" at 3,60 size 449x17
      Visibility <- "HMI Data: Warehouse HMI_screenNumber"
   Rectangle "Settings Border Hide" at 455,60 size 456x18
      Visibility <- "HMI Data: Warehouse HMI_screenNumber"
   Rectangle "Network Health Border Hide" at 914,60 size 449x18
      Visibility <- "HMI Data: Warehouse HMI_screenNumber"
   Button "Part Call Screen" at 0,0 size 455x68; TextOff 'PART CALL'
      on Release: ActivateScreen("1 PART CALL", 0)
   Button "Settings Screen" at 455,0 size 460x68; TextOff 'SETTINGS'
      on Release: ActivateScreen("2 SETTINGS", 0)
   Button "Network Health Screen" at 914,0 size 452x68; TextOff 'NW HEALTH'
   ScreenModuleView "pbSelectStation" at 60,108 size 370x55; Guid_{11997190-63616} 'Select Station'; ScreenModuleType ""
      on Guid_{11997190-211461}: function_efd93a16("Select Station", 30, 78, 1, -1, 1)
      Guid_{11997190-63605} <- "HMI Data: Warehouse HMI_settings_selectStation"
   ScreenModuleView "pbSelectWIP" at 60,173 size 370x56; Guid_{11997190-63616} 'Select WIP'; ScreenModuleType ""
      on Guid_{11997190-211461}: function_efd93a16("Select WIP", 30, 78, 1, -1, 1)
      Guid_{11997190-63605} <- "HMI Data: Warehouse HMI_settings_selectWip"
   ScreenModuleView "pbSelectButton" at 60,239 size 370x55; Guid_{11997190-63616} 'Select Button'; ScreenModuleType ""
      on Guid_{11997190-211461}: function_efd93a16("Select Button", 30, 78, 1, -1, 1)
      Guid_{11997190-63605} <- "HMI Data: Warehouse HMI_settings_selectButton"
   ScreenModuleView "pbAssign" at 60,652 size 370x56; Guid_{11997190-63616} 'Assign'; ScreenModuleType ""
      Guid_{11997190-63605} <- "HMI Data: Warehouse HMI_settings_assign"
   ScreenModuleView "iofLine" at 60,290 size 178x111; Guid_{11997190-206093} 'Line:'; ScreenModuleType ""
      Guid_{11997190-63113} <- "HMI Data: Warehouse HMI_settings_line"
   ScreenModuleView "iofDropzone" at 252,290 size 178x111; Guid_{11997190-206093} 'Dropzone:'; ScreenModuleType ""
      Guid_{11997190-63113} <- "HMI Data: Warehouse HMI_settings_dropzone"
   ScreenModuleView "iofAllotted" at 60,405 size 178x111; Guid_{11997190-206093} 'Total:'; ScreenModuleType ""
      Guid_{11997190-63113} <- "HMI Data: Warehouse HMI_settings_total"
   ScreenModuleView "iofCritical" at 252,405 size 178x111; Guid_{11997190-206093} 'Critical:'; ScreenModuleType ""
      Guid_{11997190-63113} <- "HMI Data: Warehouse HMI_settings_critical"
   TextField "tfHeaderLine" at 520,108 size 135x40; Text 'LINE'
   TextField "tfHeaderDropzone" at 655,108 size 40x40; Text 'DZ'
   TextField "tfHeaderWIP" at 695,108 size 40x40; Text 'WIP'
   TextField "tfHeaderButtonNumber" at 735,108 size 40x40; Text 'BTN'
   TextField "tfHeaderTotal" at 775,108 size 80x40; Text 'TOTAL'
   TextField "tfHeaderCritical" at 855,108 size 80x40; Text 'CRITICAL'
   TextField "tfHeaderPartNumber" at 935,108 size 256x40; Text 'PART NUMBER'
   ScreenModuleView "Settings Station Row_1" at 520,158 size 671x180; ScreenModuleType ""
      Guid_{11997190-213063} <- "HMI Data: Warehouse HMI_settings_stationRows{0}"
   ScreenModuleView "Settings Station Row_2" at 520,343 size 671x180; ScreenModuleType ""
      Guid_{11997190-213063} <- "HMI Data: Warehouse HMI_settings_stationRows{1}"
   ScreenModuleView "Settings Station Row_3" at 520,528 size 671x180; ScreenModuleType ""
      Guid_{11997190-213063} <- "HMI Data: Warehouse HMI_settings_stationRows{2}"
   ScreenModuleView "Settings Vertical Table Navigation" at 1206,108 size 100x600; ScreenModuleType ""
      Guid_{11997190-209443} <- "HMI Data: Warehouse HMI_settings_stnTableNavBar_hmi"
   ScreenModuleView "Part_Number_Entry" at 60,526 size 370x111; ScreenModuleType ""
      Guid_{11997190-63113} <- "HMI Data: Warehouse HMI_settings_partNumber"

